REGION Network 1 (SCL)
   //---------------------------------------------------------------------
   //In this network first, we assign the ip address and port number for the printer (MarkemImaje). Then prepare the command for 
   //time synch, checking alarms, sending a batch number, intiating counter and selecting the label. one port for all data.
   //---------------------------------------------------------------------
   //
   REGION AddressAssign
       (*
       //Special case: if ip and port is entered correctly but still the communication not established, try onece more.
       IF #ConnectionStatus = False AND #ErrorIP = FALSE AND #ReTry = FALSE AND #ConnAgainT.Q = FALSE AND #TimeOutError = FALSE THEN
           #ReTry := True;
       ELSE
           #ReTry := FALSE;
       END_IF;
       *)
       // ip and port assign to the printer
       #Config := "LGF_StringToTaddr"(ipAddressString := #RemoteAddress, error => #ErrorIP, status => #StatusIP);
       //when IP address change, disconnect and connect again
       #ChangeIP_T(IN:=#RemoteAddressOld <> #RemoteAddress,
                   PT:=T#2S);
       IF #ChangeIP_T.Q OR #ErrorIP = TRUE THEN
           #IP_Change := TRUE;
       ELSE
           #IP_Change := FALSE;
       END_IF;
       #RemoteAddressOld := #RemoteAddress;
       FOR #i := 1 TO 4 DO
           #Configuration.connection.partnerIP.ADDR[#i] := USINT_TO_BYTE(#Config.REM_IP_ADDR[#i]);//assign ip address
       END_FOR;
       //assign id port and other setting for TCP communication
       #Configuration.connection.connectionID := #ID;
       #Configuration.connection.comService := 1;
       //if it is active connection
       IF #ConType = TRUE THEN
           #Configuration.connection.isClient := True;
           IF #Config.REM_PORT_NR = 0 THEN
               #Configuration.connection.partnerPort := 9100; // default port for Markem communication
           ELSE
               #Configuration.connection.partnerPort := #Config.REM_PORT_NR;
           END_IF;
       ELSE //if it is passive connection
           #Configuration.connection.isClient := FALSE;
           #Configuration.connection.localPort := 2000;
       END_IF;
   END_REGION
   REGION HMI
       // Data for the HMI
       #DatePrinted := DELETE(IN:=#Date, L:=2, P:=1);
       #TimePrinted := DELETE(IN := #Time, L := 2, P := 5);
       #TimePrinted := INSERT(IN1 := #TimePrinted, IN2 := ':', P := 2);
       IF #ExtDate <> '' THEN
           #ExpFlag := TRUE;
       ELSE
           #ExpFlag := FALSE;
       END_IF;
   END_REGION

   REGION Commands 
       // Creating Commands and preparing them to Send
       IF #Step = 1 THEN
           //command for time synchronisation
           #CommandHead := 'V21'; //head for time/date synch
           #SData[0] := #Start;
           Strg_TO_Chars(Strg := #CommandHead,
                         pChars := 1,
                         Cnt => #Dummy2,
                         Chars := #SData);
           #SData[4] := ' ';
           Strg_TO_Chars(Strg := #Date,
                         pChars := 0,
                         Cnt => #Dummy2,
                         Chars := #DateChar);
           FOR #i := 5 TO 8 DO
               #SData[#i] := #DateChar[#i - 5];
           END_FOR;
           #SData[9] := '-';
           #SData[10] := #DateChar[4];
           #SData[11] := #DateChar[5];
           #SData[12] := '-';
           #SData[13] := #DateChar[6];
           #SData[14] := #DateChar[7];
           #SData[15] := #NewLine;
           //sending time
           #SData[16] := #Start;
           #SData[17] := 'V';
           #SData[18] := '2';
           #SData[19] := '0';
           #SData[20] := ' ';
           Strg_TO_Chars(Strg := #Time,
                         pChars := 0,
                         Cnt => #Dummy2,
                         Chars := #TimeChar);
           #SData[21] := #TimeChar[0];
           #SData[22] := #TimeChar[1];
           #SData[23] := ':';
           #SData[24] := #TimeChar[2];
           #SData[25] := #TimeChar[3];
           #SData[26] := ':';
           #SData[27] := #TimeChar[4];
           #SData[28] := #TimeChar[5];
           #SData[29] := #End;
           #RLen := 2;
           #SLen := 30;
           #Step := 0;
           #STrig := TRUE;
           #RdataTime := TRUE;
           #RdataAlarm := FALSE;
           #RdataBatch := FALSE;
           #RdataMacro := FALSE;
       ELSIF #Step = 2 THEN
           //command for checking the alarms
           #CommandHead := 'S100'; //head for current status of the printer
           #SData[0] := #Start;
           Strg_TO_Chars(Strg := #CommandHead,
                         pChars := 1,
                         Cnt => #Dummy2,
                         Chars := #SData);
           #SData[5] := #End;
           #RLen := 34;
           #SLen := 6;
           #STrig := TRUE;
           #Step := 0;
           #RdataAlarm := TRUE;
           #RdataTime := FALSE;
           #RdataBatch := FALSE;
           #RdataMacro := FALSE;
       ELSIF #Step = 3 THEN
           //command for sending variable text
           #SData[0] := #Start;
           #CommandHead := 'W1 "';
           //GTIN number 14 digits
           Strg_TO_Chars(Strg := #CommandHead,
                         pChars := 1,
                         Cnt => #Dummy2,
                         Chars := #SData);
           Strg_TO_Chars(Strg := #GTIN_Number,
                         pChars := 5,
                         Cnt => #Dummy2,
                         Chars := #SData);
           #SData[19] := '"';
           #SData[20] := #NewLine;
           //Batch
           #CommandHead := '!W4 "';
           //Batch number 10 digits
           Strg_TO_Chars(Strg := #CommandHead,
                         pChars := 21,
                         Cnt => #Dummy2,
                         Chars := #SData);
           Strg_TO_Chars(Strg := #BatchNumber,
                         pChars := 26,
                         Cnt => #Dummy2,
                         Chars := #SData);
           #SData[36] := '"';
           #SData[37] := #NewLine;
           //Article number
           #CommandHead := '!W5 "';
           //Article number 10 digits
           Strg_TO_Chars(Strg := #CommandHead,
                         pChars := 38,
                         Cnt => #Dummy2,
                         Chars := #SData);
           Strg_TO_Chars(Strg := #ArtNumber,
                         pChars := 43,
                         Cnt => #Dummy2,
                         Chars := #SData);
           #SData[53] := '"';
           #SData[54] := #NewLine;
           //Ext date
           #CommandHead := '!W3 "';
           //Ext date 6 digits
           Strg_TO_Chars(Strg := #CommandHead,
                         pChars := 55,
                         Cnt => #Dummy2,
                         Chars := #SData);
           IF #ExtDate <> '' THEN //if expiration date is available 
               Strg_TO_Chars(Strg := #ExtDate,
                             pChars := 60,
                             Cnt => #Dummy2,
                             Chars := #SData);
           ELSE
               FOR #i := 60  TO 65 DO
                   #SData[#i] := ' ';
               END_FOR;
           END_IF;
           #SData[66] := '"';
           #SData[67] := #NewLine;
           //Machine ID
           #CommandHead := '!W6 "';
           //Machine ID 3 digits
           Strg_TO_Chars(Strg := #CommandHead,
                         pChars := 68,
                         Cnt => #Dummy2,
                         Chars := #SData);
           Strg_TO_Chars(Strg := #MachineID,
                         pChars := 73,
                         Cnt => #Dummy2,
                         Chars := #SData);
           //Reinit the counter 
           #SData[76] := '"';
           #SData[77] := #NewLine;
           VAL_STRG(IN := (#Serial+1),// +1 to make sure we have no TRP with same serial
                    SIZE := 0,
                    PREC := 0,
                    FORMAT := 0,
                    P := 1,
                    OUT => #SerialSTR);
           #SerialLen := LEN(#SerialSTR);
           #CommandHead := '!N1 ';//!N1 "Serial" 1 5 1
           Strg_TO_Chars(Strg := #CommandHead,
                         pChars := 78,
                         Cnt => #Dummy2,
                         Chars := #SData);
           #CommandHead := #SerialSTR;
           Strg_TO_Chars(Strg := #CommandHead,
                         pChars := 82,
                         Cnt => #Dummy2,
                         Chars := #SData);
           #CommandHead := ' 1 5 1';
           Strg_TO_Chars(Strg := #CommandHead,
                         pChars := 82+#SerialLen,
                         Cnt => #Dummy2,
                         Chars := #SData);
           #SData[82 + #SerialLen + 6] := #End;
           #RLen := 0;
           #SLen := INT_TO_UDINT( 82 + #SerialLen + 6 + 1);
           #Step := 0;
           #STrig := TRUE;
           #Selected := FALSE;
           #RdataTime := FALSE;
           #RdataAlarm := FALSE;
           #RdataBatch := TRUE;
           #RdataMacro := FALSE;
       //command for selectiong the Macro 
       ELSIF #Step = 4 THEN
           #CommandHead := 'M "'; //head for selecting the Macro
           #SData[0] := #Start;
           Strg_TO_Chars(Strg := #CommandHead,
                         pChars := 1,
                         Cnt => #Dummy2,
                         Chars := #SData);
           IF #ExtDate = '' THEN
               IF #Inverse = TRUE THEN
                   Strg_TO_Chars(Strg := #LabelNameInv,
                                 pChars := 4,
                                 Cnt => #Dummy2,
                                 Chars := #SData);
               ELSE
                   Strg_TO_Chars(Strg := #LabelName,
                                 pChars := 4,
                                 Cnt => #Dummy2,
                                 Chars := #SData);
               END_IF;
           ELSE
               IF #Inverse = TRUE THEN
                   Strg_TO_Chars(Strg := #LabelNameExpInv,
                                 pChars := 4,
                                 Cnt => #Dummy2,
                                 Chars := #SData);
               ELSE
                   Strg_TO_Chars(Strg := #LabelNameExp,
                                 pChars := 4,
                                 Cnt => #Dummy2,
                                 Chars := #SData);
               END_IF;
           END_IF;
           #SData[16] := '"';
           #SData[17] := #NewLine;
           IF #Stop = TRUE THEN
               #SData[18] := ' ';
               #SData[19] := 'p';
           ELSE
               #SData[18] := #Start;
               #SData[19] := 'p';
           END_IF;
           #SData[20] := #End;
           #RLen := 2;
           #SLen := 21;
           #Step := 0;
           #STrig := TRUE;
           #RdataTime := FALSE;
           #RdataAlarm := FALSE;
           #RdataBatch := FALSE;
           #RdataMacro := TRUE;
       ELSE
           #STrig := FALSE;
       END_IF;
   END_REGION

   REGION Feedback
       // Statement section REGION
       //Expect to receive "ACT"
       IF #DataReceived = TRUE THEN
           #StartTNR := FALSE;
           IF #RdataTime = TRUE THEN //check for the feedback for the time command
               FOR #i := 0 TO 56 DO
                   #TimeReceivedData[#i] := #RData[#i];
               END_FOR;
               IF #TimeReceivedData[0] = #NewLine THEN
                   #TimeOK := TRUE;
                   #TimeReceivedData[0] := 16#30;//clear the buffer
               ELSE
                   #TimeOK := FALSE;
               END_IF;
               #RdataTime := FALSE; // make the flag false
           ELSIF #RdataAlarm = TRUE THEN//check for the feedback for the alarm command
               FOR #i := 0 TO 56 DO
                   #AlarmReceivedData[#i] := #RData[#i];
               END_FOR;
               IF #AlarmReceivedData[32] = #End THEN // the plc receives the responce
                   #AlarmCheck := TRUE;
                   #AlarmReceivedData[32] := 16#30;//clear the buffer
                   FOR #i := 0 TO 31 DO//save the status data for processing
                       IF #AlarmReceivedData[#i] = '1' THEN
                           #PrinterAlarmStatus[#i] := TRUE;
                       ELSE
                           #PrinterAlarmStatus[#i] := FALSE;
                       END_IF;
                   END_FOR;
               ELSE
                   #AlarmCheck := FALSE;
               END_IF;
               #RdataAlarm := FALSE;
           //ELSIF #RdataBatch = TRUE THEN //no feedback from the command except batch
               //         FOR #i := 0 TO 56 DO
               //            #BatchReceivedData[#i] := #RData[#i];
               //        END_FOR;
               //       IF #BatchReceivedData[0] = 16#24 THEN
             //  #BatchOK := TRUE;
               //           #BatchReceivedData[0] := 16#30;//clear the buffer
               //       ELSE
               //        #BatchOK := FALSE;
               //    END_IF;
               //     #RdataBatch := FALSE;
           ELSIF #RdataMacro = TRUE OR #RdataBatch = TRUE THEN
               FOR #i := 0 TO 56 DO
                   #MacroReceivedData[#i] := #RData[#i];
               END_FOR;
               IF #MacroReceivedData[0] = #NewLine THEN // the plc receives the responce
                   #LabelOK := TRUE;
                   #MacroReceivedData[0] := 16#30;//clear the buffer
               ELSE
                   #LabelOK := FALSE;
               END_IF;
               #RdataMacro := FALSE;
           END_IF;
       ELSIF #DataSent = TRUE AND #RdataAlarm = TRUE OR #RdataTime = TRUE OR #RdataMacro = TRUE THEN // command send noting received
           #StartTNR := TRUE;
           IF #RdataTime = TRUE THEN
               #TimeOK := FALSE;
           END_IF;
           IF #RdataAlarm = TRUE THEN
               #AlarmCheck := FALSE;
           END_IF;
           IF #RdataMacro = TRUE THEN
               #LabelOK := FALSE;
           END_IF;
       END_IF;
   END_REGION

   REGION Sending
       //selecting the label properties for every instalation of the new printer or power OFF then ON
       #SelectingR(CLK:=#LabelSelecting);
       #ReconnectR(CLK := #ConnectionStatus);
       #InverseR(CLK:=#Inverse);
       #InverseF(CLK:=#Inverse);
        // it is assumed at every reconnection the label is gone so, we send it again
       IF #SelectingR.Q = TRUE OR #ReconnectR.Q = TRUE OR #InverseR.Q = TRUE OR #InverseF.Q = TRUE THEN
           #Step := 4;
           #Selected := TRUE;
       END_IF;
       // set the step to 3 after label is selecting (small delay to make sure that the label is loaded)
       #BatchAfterLabelT(IN := #Selected,
                         PT := T#5S);
       IF #BatchAfterLabelT.Q = TRUE THEN
           #Step := 3;
       END_IF;
       // Send the updateble data when it is changed and step 4 is done
       IF #PlainDataChanged = TRUE AND #SelectingR.Q = FALSE THEN
           #Step := 3;
           #Selected := FALSE;
       END_IF;
       // Send time and alarm commands
       //every 10 minute synchronise time
       #TimeSynchT(IN := #TimeSynchEnable,
                  PT := #TimeSynchPeriod);
       IF #TimeSynchT.Q = TRUE THEN
           #Step := 1;
           #TimeSynchEnable := FALSE;
       ELSIF #ConnectionStatus = TRUE AND NOT (#SelectingR.Q = TRUE OR #ReconnectR.Q = TRUE OR #InverseR.Q = TRUE OR #InverseF.Q = TRUE) AND #PlainDataChanged = FALSE THEN
           #TimeSynchEnable := True;
       ELSE
           #TimeSynchEnable := FALSE;
       END_IF;
       //every 5 minute check for alarm
       #AlarmCheckT(IN := #AlarmCheckEnable,
                   PT := #AlarmCheckPeriod + T#20MS);//+20ms to avoid conflict
       IF #AlarmCheckT.Q = TRUE THEN
           #Step := 2;
           #AlarmCheckEnable := FALSE;
       ELSIF #ConnectionStatus = TRUE AND NOT (#SelectingR.Q = TRUE OR #ReconnectR.Q = TRUE OR #InverseR.Q = TRUE OR #InverseF.Q = TRUE) AND #PlainDataChanged = FALSE THEN
           #AlarmCheckEnable := TRUE;
       ELSE
           #AlarmCheckEnable := FALSE;
       END_IF;
   END_REGION
   (*
   REGION ConnReestablised
       // connection Re-Established Rotinue. It try 5 times to connect to the printer, if not succsess enable time out error
       #ConnAgainT(IN := #ReTry,
                  PT := T#5S);// time out for reconnection
       //try five times to connect
       #ConnTryCountC(CU := #ReTry,
                     R := #ConnectionStatus,
                     PV := 5,
                     Q => #TimeOutError);
   END_REGION
   *)
   REGION send try
       //if not receiving feedback after 10ms send a commad again
       #NotReceiveT(IN := #StartTNR,
                   PT := #TimeNR,
                   Q => #SendAgainTrigger);
       IF #SendAgainTrigger = TRUE THEN
           #StartTNR := FALSE;
       END_IF;
    //   #NotReceivingError(IN:= NOT(#TimeOK AND #LabelOK AND #NoAlarm = FALSE), // if we are not receiving a feedback after sending two times pop up an alarm
    //                      PT:=T#90S,
    //                      Q=>#CommandError);
   END_REGION

   REGION Counter
       // count the number of the trigger and initiated it when sending the label information. the counter only restarted when the batch changed. 
       #ExtTriggerR(CLK:=#ExtTrigger);
       IF #ExtTriggerR.Q = TRUE THEN
           "Counter_32Bit_1"(Varia := 1,
                           CountedValue := #Serial);
       END_IF;
       IF #Serial > 99999 OR #PlainDataChanged = TRUE THEN //restart the counter if it reaches the limit or data changed at Plain
           #Serial := 0;
       END_IF;
   END_REGION
END_REGION
END_FUNCTION_BLOCK

FUNCTION_BLOCK "Domino_AX"   // FB6, LAD
{ S7_Optimized_Access := 'TRUE' }
VERSION : 0.1
   VAR_INPUT
      RemoteAddress : String[20];
      ConnectionStatus : Bool;
      ID : Conn_Ouc;
      ConType : Bool;
      ArtFlag : Bool;
      MDR_Flag : Bool;
      BatchStatus : USInt;
      BatchNumber : String;
      ArtBaseNumber : String;
      MarketRegCode : String;
      ExtDate : String;
      "Date" : String;
      "Time" : String;
      PlainDataChanged : Bool;
      DataReceived : Bool;
      DataReceivedBatch : Bool;
      DataSent : Bool;
      DataSentBatch : Bool;
      TimeSynchPeriod : Time := T#10M;
      AlarmCheckPeriod : Time := T#5M;
      RDataBatch : Array[0..56] of Byte;
      RData : Array[0..56] of Byte;
      NMDR_LabelName : String;
      LabelSelecting : Bool;
   END_VAR
   VAR_OUTPUT
      ErrorIP : Bool;
      BatchOK : Bool;
      AlarmCheck : Bool;
      TimeOK : Bool;
      LabelOK : Bool;
   END_VAR
   VAR
      Config : TADDR_Param;
      Configuration : "typeLCom_Config";
      ConfigurationBatch : "typeLCom_Config";
      RLen : UDInt;
      RLenMDR : UDInt;
      SLen : UDInt;
      SLenMDR : UDInt;
      SData : Array[0..56] of Byte;
      SDataMDR : Array[0..99] of Byte;
      StartTNRMDR : Bool;
      StartTNR : Bool;
      TimeNR : Time := T#1m;
      SendAgainTrigger : Bool;
      SendAgainTriggerBatch : Bool;
      NotReceiveT : TON_TIME;
      NotReceiveBatchT : TON_TIME;
      TimeSynchEnable : Bool := false;
      TimeSynchT : TON_TIME;
      AlarmCheckEnable : Bool := false;
      AlarmCheckT : TON_TIME;
      STrig : Bool;
      StrigBatch : Bool;
      "Step" : UDInt;
      AlarmReceivedData : Array[0..56] of Byte;
      TimeReceivedData : Array[0..56] of Byte;
      BatchReceivedData : Array[0..56] of Byte;
      LabelReceivedData : Array[0..56] of Byte;
      PrinterAlarmStatus : Array[0..8] of Char;
      RdataTime : Bool;
      RdataAlarm : Bool;
      RdataLabel : Bool;
      BlockedProduct : Bool;
      SelectingR : R_TRIG;
      Selected : Bool;
      ReconnectR : R_TRIG;
      MDR_R : R_TRIG;
      MDR_F : F_TRIG;
      BlockedR : R_TRIG;
      BlockedF : F_TRIG;
      ActualNMDR_Label : String;
      NLabelChanged : Bool;
      BatchAfterLabelT : TON_TIME;
      ChangeIP_T : TP_TIME;
      IP_Change : Bool;
      RemoteAddressOld : String;
   END_VAR
   VAR_TEMP
      StatusIP : Word;
      Dummy2 : UInt;
      i : Int;
      CommandHead : String;
      SecondRowSTR : String;
      SecondRowSTR1 : String;
      LenDummy : Int;
      ArtLen : Int;
      LenLabel : Int;
      LenLabelSTR : String;
      LabelCommand : String;
   END_VAR
   VAR CONSTANT
      Start : Char := '$1B';
      Start1 : Char := '$02';
      End1 : Char := '$03';
      End : Char := '$04';
      MDR_LabelName1 : String := 'MDR1';
      MDR_LabelName2 : String := 'MDR2';
   END_VAR
BEGIN

REGION Network 1 (SCL)
   //---------------------------------------------------------------------
   //In this network first, we assign the ip address and port number for the printer (Domino_AX). Then prepare the command for 
   //time synch, receiving alarms and sending a batch number. one port (16000) for the batch number and another port for the rest.
   //---------------------------------------------------------------------
   REGION Address_Assign
       (*
       //Special case: if ip and port is entered correctly but still the communication not established, try onece more.
       IF #ConnectionStatus = False AND #ErrorIP = FALSE AND #ReTry = FALSE AND #ConnAgainT.Q = FALSE AND #TimeOutError = FALSE THEN
           #ReTry := True;
       ELSE
           #ReTry := FALSE;
       END_IF;
       *)
       // ip and port assign to the printer
       #Config := "LGF_StringToTaddr"(ipAddressString := #RemoteAddress, error => #ErrorIP, status => #StatusIP);
       //when IP address change, disconnect and connect again
       #ChangeIP_T(IN := #RemoteAddressOld <> #RemoteAddress,
                   PT := T#2S);
       IF #ChangeIP_T.Q OR #ErrorIP = TRUE THEN
           #IP_Change := TRUE;
       ELSE
           #IP_Change := FALSE;
       END_IF;
       #RemoteAddressOld := #RemoteAddress;
       FOR #i := 1 TO 4 DO
          #Configuration.connection.partnerIP.ADDR[#i] := USINT_TO_BYTE(#Config.REM_IP_ADDR[#i]);//assign ip address
          #ConfigurationBatch.connection.partnerIP.ADDR[#i] := USINT_TO_BYTE(#Config.REM_IP_ADDR[#i]);//assign ip address
      END_FOR;

       //assign id port and other setting for TCP communication
       #Configuration.connection.connectionID := #ID;
       #Configuration.connection.comService := 1;
       #ConfigurationBatch.connection.connectionID := #ID + 1;
       #ConfigurationBatch.connection.comService := 1;
       #ConfigurationBatch.connection.isClient := True;
       #ConfigurationBatch.connection.partnerPort := 16000;// only for domino printer
         //if it is active connection
       IF #ConType = TRUE THEN
           #Configuration.connection.isClient := True;
           IF #Config.REM_PORT_NR = 0 THEN
               #Configuration.connection.partnerPort := 7000; // default port for domino communication
           ELSE
               #Configuration.connection.partnerPort := #Config.REM_PORT_NR;
           END_IF;
       ELSE //if it is passive connection
           #Configuration.connection.isClient := FALSE;
           #Configuration.connection.localPort := 2000;
       END_IF;

   END_REGION
   REGION Trigger
       // Trigger signal to send a correct data for print when Batch ended
       IF #BatchStatus = 3 THEN
           #BlockedProduct := TRUE;
       ELSE
           #BlockedProduct := FALSE;
       END_IF;
       // Trigger signal to send Non-MDR label when it is changed from the screen
       IF #MDR_Flag = FALSE AND #ActualNMDR_Label <> #NMDR_LabelName THEN
           #NLabelChanged := TRUE;
           #ActualNMDR_Label := #NMDR_LabelName;
       ELSE
           #NLabelChanged := FALSE;
       END_IF;
   END_REGION

   REGION Commands
         //command for time synchronisation
         IF #Step = 1 THEN
             #CommandHead := 'C'; //head for time
             #SData[0] := #Start;
             Strg_TO_Chars(Strg := #CommandHead,
                           pChars := 1,
                           Cnt => #Dummy2,
                           Chars := #SData);
             Strg_TO_Chars(Strg := #Date,
                           pChars := 2,
                           Cnt => #Dummy2,
                           Chars := #SData);
             #SData[10] := '0';
             #SData[11] := '0';
             Strg_TO_Chars(Strg := #Time,
                           pChars := 12,
                           Cnt => #Dummy2,
                           Chars := #SData);
             #SData[18] := #End;
             #RLen := 1;
             #SLen := 19;
             #STrig := TRUE;
             #Step := 0; //idea state
             #RdataTime := TRUE;
             #RdataAlarm := FALSE;
             #RdataLabel := FALSE;

         ELSIF #Step = 2 THEN
             //command for checking the alarms
             #CommandHead := 'O1?'; //head for current status of the printer
             #SData[0] := #Start;
             Strg_TO_Chars(Strg := #CommandHead,
                           pChars := 1,
                           Cnt => #Dummy2,
                           Chars := #SData);
             #SData[4] := #End;
             #RLen := 9;
             #SLen := 5;
             #STrig := TRUE;
             #Step := 0; 
             #RdataAlarm := TRUE;
             #RdataTime := FALSE;
             #RdataLabel := FALSE;
             (*  we should creat a MDR layout at the Printer with two fields. one id used for batch+art base and the 
                   second is use for market Reg and Ext date*)
                   //Constructiong the buffer command in the first row
         ELSIF #Step=3 THEN
             #RLenMDR := 1; // receive 0x06 as an acknowledgment
             #StrigBatch := TRUE;
             #Step := 0;
             #Selected := FALSE;
                 #SDataMDR[0] := #Start1;
                 Strg_TO_Chars(Strg := #BatchNumber,
                               pChars := 1,
                               Cnt => #Dummy2,
                               Chars := #SDataMDR);
                 IF #ArtFlag = TRUE AND #MarketRegCode <> '' AND #ExtDate <> '' THEN // print all information in two rows
                     #SDataMDR[11] := ' '; //space
                     #SDataMDR[12] := 'A';
                     #SDataMDR[13] := 'R';
                     #SDataMDR[14] := 'T';
                     #ArtLen := LEN(#ArtBaseNumber);
                     Strg_TO_Chars(Strg := #ArtBaseNumber,
                                   pChars := 15,
                                   Cnt => #Dummy2,
                                   Chars := #SDataMDR);
                     IF #BatchStatus = 3 THEN //add a sign '+' at the con
                         #SDataMDR[15 + #ArtLen] := '+';

                     ELSE
                         #SDataMDR[15 + #ArtLen] := ' ';
                     END_IF;
                     #SDataMDR[15 + #ArtLen + 1] := ',';//seprator for the second row
                     #SecondRowSTR := CONCAT(IN1 := #MarketRegCode, IN2 := 'BBD');
                     #SecondRowSTR1 := CONCAT(IN1 := #SecondRowSTR, IN2 := #ExtDate);
                     #LenDummy := LEN(#SecondRowSTR1);
                     Strg_TO_Chars(Strg := #SecondRowSTR1,
                                   pChars := 15 + #ArtLen + 2,
                                   Cnt => #Dummy2,
                                   Chars := #SDataMDR);
                     #SDataMDR[15 + #ArtLen + 2 + #LenDummy] := #End1;
                     #SLenMDR := 15 + #ArtLen + 2 + #LenDummy + 1;
                 ELSIF #ArtFlag = TRUE AND #MarketRegCode <> '' AND #ExtDate = '' THEN // print all information exept expiration date in two rows
                     #SDataMDR[11] := ' '; //space
                     #SDataMDR[12] := 'A';
                     #SDataMDR[13] := 'R';
                     #SDataMDR[14] := 'T';
                     #ArtLen := LEN(#ArtBaseNumber);
                     Strg_TO_Chars(Strg := #ArtBaseNumber,
                                   pChars := 15,
                                   Cnt => #Dummy2,
                                   Chars := #SDataMDR);
                     IF #BatchStatus = 3 THEN //add a sign '+' at the con
                         #SDataMDR[15 + #ArtLen] := '+';

                     ELSE
                         #SDataMDR[15 + #ArtLen] := ' ';
                     END_IF;
                     #SDataMDR[15 + #ArtLen + 1] := ',';//seprator for the second row
                     #LenDummy := LEN(#MarketRegCode);
                     Strg_TO_Chars(Strg := #MarketRegCode,
                                   pChars := 15 + #ArtLen + 2,
                                   Cnt => #Dummy2,
                                   Chars := #SDataMDR);
                     #SDataMDR[15 + #ArtLen + 2 + #LenDummy] := #End1;
                     #SLenMDR := 15 + #ArtLen + 2 + #LenDummy + 1;
                 ELSIF #ArtFlag = TRUE AND #MarketRegCode = '' AND #ExtDate <> '' THEN // print all information exept Market reg code in two rows
                     #SDataMDR[11] := ' '; //space
                     #SDataMDR[12] := 'A';
                     #SDataMDR[13] := 'R';
                     #SDataMDR[14] := 'T';
                     #ArtLen := LEN(#ArtBaseNumber);
                     Strg_TO_Chars(Strg := #ArtBaseNumber,
                                   pChars := 15,
                                   Cnt => #Dummy2,
                                   Chars := #SDataMDR);
                     IF #BatchStatus = 3 THEN //add a sign '+' at the con
                         #SDataMDR[15 + #ArtLen] := '+';

                     ELSE
                         #SDataMDR[15 + #ArtLen] := ' ';
                     END_IF;
                     #SDataMDR[15 + #ArtLen + 1] := ',';//seprator for the second row
                     #SecondRowSTR1 := CONCAT(IN1 := 'BBD', IN2 := #ExtDate);
                     #LenDummy := LEN(#SecondRowSTR1);
                     Strg_TO_Chars(Strg := #SecondRowSTR1,
                                   pChars := 15 + #ArtLen + 2,
                                   Cnt => #Dummy2,
                                   Chars := #SDataMDR);
                     #SDataMDR[15 + #ArtLen + 2 + #LenDummy] := #End1;
                     #SLenMDR := 15 + #ArtLen + 2 + #LenDummy + 1;
                 ELSIF #ArtFlag = TRUE AND #MarketRegCode = '' AND #ExtDate = '' THEN // print only in one row
                     #SDataMDR[11] := ' '; //space
                     #SDataMDR[12] := 'A';
                     #SDataMDR[13] := 'R';
                     #SDataMDR[14] := 'T';
                     #ArtLen := LEN(#ArtBaseNumber);
                     Strg_TO_Chars(Strg := #ArtBaseNumber,
                                   pChars := 15,
                                   Cnt => #Dummy2,
                                   Chars := #SDataMDR);
                     IF #BatchStatus = 3 THEN //add a sign '+' at the con
                         #SDataMDR[15 + #ArtLen] := '+';

                     ELSE
                         #SDataMDR[15 + #ArtLen] := ' ';
                     END_IF;
                     #SDataMDR[16 + #ArtLen] := #End1;
                     #SLenMDR := 16 + #ArtLen + 1;
                 ELSIF #ArtFlag = FALSE AND #MarketRegCode <> '' AND #ExtDate <> '' THEN // print all information exept art flag  in two rows
                     IF #BatchStatus = 3 THEN //add a sign '+' at the con
                         #SDataMDR[11] := '+';

                     ELSE
                         #SDataMDR[11] := ' ';
                     END_IF;
                     #SDataMDR[12] := ',';//seprator for the second row
                     #SecondRowSTR := CONCAT(IN1 := #MarketRegCode, IN2 := 'BBD');
                     #SecondRowSTR1 := CONCAT(IN1 := #SecondRowSTR, IN2 := #ExtDate);
                     #LenDummy := LEN(#SecondRowSTR1);
                     Strg_TO_Chars(Strg := #SecondRowSTR1,
                                   pChars := 13,
                                   Cnt => #Dummy2,
                                   Chars := #SDataMDR);
                     #SDataMDR[13 + #LenDummy] := #End1;
                     #SLenMDR := 13 + #LenDummy + 1;
                 ELSIF #ArtFlag = FALSE AND #MarketRegCode <> '' AND #ExtDate = '' THEN // print all information exept expiration art number and ext date in two rows
                     IF #BatchStatus = 3 THEN //add a sign '+' at the con
                         #SDataMDR[11] := '+';

                     ELSE
                         #SDataMDR[11] := ' ';
                     END_IF;
                     #SDataMDR[12] := ',';//seprator for the second row
                     #LenDummy := LEN(#MarketRegCode);
                     Strg_TO_Chars(Strg := #MarketRegCode,
                                   pChars := 13,
                                   Cnt => #Dummy2,
                                   Chars := #SDataMDR);
                     #SDataMDR[13 + #LenDummy] := #End1;
                     #SLenMDR := 13 + #LenDummy + 1;
                 ELSIF #ArtFlag = FALSE AND #MarketRegCode = '' AND #ExtDate <> '' THEN // print in one row
                     IF #BatchStatus = 3 THEN //add a sign '+' at the con
                         #SDataMDR[11] := '+';

                     ELSE
                         #SDataMDR[11] := ' ';
                     END_IF;
                     #SDataMDR[12] := ',';//seprator for the second row
                     #SecondRowSTR1 := CONCAT(IN1 := 'BBD', IN2 := #ExtDate);
                     #LenDummy := LEN(#SecondRowSTR1);
                     Strg_TO_Chars(Strg := #SecondRowSTR1,
                                   pChars := 13,
                                   Cnt => #Dummy2,
                                   Chars := #SDataMDR);
                     #SDataMDR[13 + #LenDummy] := #End1;
                     #SLenMDR := 13 + #LenDummy + 1;
                 ELSE // print only batch
                     IF #BatchStatus = 3 THEN //add a sign '+' at the con
                         #SDataMDR[11] := '+';

                     ELSE
                         #SDataMDR[11] := ' ';
                     END_IF;
                     #SDataMDR[12] := #End1;
                     #SLenMDR := 13;
                 END_IF;
         ELSIF #Step =4 THEN
             //command for selecting the label
             #CommandHead := 'ON1'; //head for current status of the printer
             #SData[0] := #Start;
             Strg_TO_Chars(Strg := #CommandHead,
                           pChars := 1,
                           Cnt => #Dummy2,
                           Chars := #SData);
             IF #MDR_Flag = TRUE THEN //select the MDR layout 
                 IF #ExtDate <> '' OR #MarketRegCode <> '' THEN
                     #LabelCommand := CONCAT(IN1 := '04', IN2 := #MDR_LabelName2);
                 ELSE
                     #LabelCommand := CONCAT(IN1 := '04', IN2 := #MDR_LabelName1);
                 END_IF;
                 Strg_TO_Chars(Strg := #LabelCommand,
                               pChars := 4,
                               Cnt => #Dummy2,
                               Chars := #SData);
                 #SData[10] := #End;
                 #RLen := 1;
                 #SLen := 11;
             ELSE
                 #LenLabel := LEN(#NMDR_LabelName);
                 VAL_STRG(IN := #LenLabel,
                          SIZE := 2,
                          PREC := 0,
                          FORMAT := 0,
                          P := 1,
                          OUT => #LenLabelSTR);
                 #LabelCommand := CONCAT(IN1 := #LenLabelSTR, IN2 := #NMDR_LabelName);

                 Strg_TO_Chars(Strg := #LabelCommand,
                               pChars := 4,
                               Cnt => #Dummy2,
                               Chars := #SData);
                 FOR #i := 4 TO 5 DO //check for null char due to size
                     IF #SData[#i] = ' ' THEN
                         #SData[#i] := '0';
                     END_IF;
                 END_FOR;
                 #SData[6 + #LenLabel] := #End;
                 #RLen := 1;
                 #SLen := 7 + #LenLabel;
             END_IF;
             #STrig := TRUE;
             #Step := 0; 
             #RdataAlarm := FALSE;
             #RdataTime := FALSE;
             #RdataLabel := TRUE;
         ELSE
             #STrig := FALSE;
             #StrigBatch := FALSE;
         END_IF;
     END_REGION
       REGION Feedback
           // Statement section REGION
           //Expect to receive "ACT"
           IF #DataReceived = TRUE THEN
               #StartTNR := FALSE;
               IF #RdataTime = TRUE THEN //check for the feedback for the time command
                   FOR #i := 0 TO 56 DO
                       #TimeReceivedData[#i] := #RData[#i];
                   END_FOR;
                   IF #TimeReceivedData[0] = 16#06 THEN
                       #TimeOK := TRUE;
                       #TimeReceivedData[0] := 16#30;//clear the buffer
                   ELSE
                       #TimeOK := FALSE;
                   END_IF;
                   #RdataTime := FALSE;

               ELSIF #RdataAlarm = TRUE THEN//check for the feedback for the alarm command
                   FOR #i := 0 TO 56 DO
                       #AlarmReceivedData[#i] := #RData[#i];
                   END_FOR;
                   IF #AlarmReceivedData[1] = 'O' AND #AlarmReceivedData[2] = '1' THEN // check the responce and save them
                       #AlarmCheck := TRUE;
                       FOR #i := 0 TO 8 DO
                           #PrinterAlarmStatus[#i] := #AlarmReceivedData[#i];//save the status data for processing
                       END_FOR;
                       #AlarmReceivedData[1] := '0';//clear the buffer
                   ELSE
                       #AlarmCheck := FALSE;
                   END_IF;
                   #RdataAlarm := FALSE;
               ELSIF #RdataLabel = TRUE THEN // check for the label command feedback
                   FOR #i := 0 TO 56 DO
                       #LabelReceivedData[#i] := #RData[#i];
                   END_FOR;
                   IF #LabelReceivedData[0] = 16#06 THEN // check the responce and save them
                       #LabelOK := TRUE;
                       #LabelReceivedData[0] := '0';//clear the buffer
                   ELSE
                       #LabelOK := FALSE;
                   END_IF;
                   #RdataLabel := FALSE;
               END_IF;
           ELSIF #DataSent = TRUE THEN // command send noting received
                   #StartTNR := TRUE;
                   IF #RdataTime = TRUE THEN
                       #TimeOK := FALSE;
                   END_IF;
                   IF #RdataAlarm = TRUE THEN
                       #AlarmCheck := FALSE;
                   END_IF;
                   IF #RdataLabel = TRUE THEN
                       #LabelOK := FALSE;
                   END_IF;
               END_IF;
               //Expect to receive "ACT" for external Info Command
               IF #DataReceivedBatch = TRUE THEN
                   #StartTNRMDR := FALSE;
                   FOR #i := 0 TO 56 DO
                       #BatchReceivedData[#i] := #RDataBatch[#i];
                   END_FOR;
                   IF #BatchReceivedData[0] = 16#06 THEN
                       #BatchOK := TRUE;
                   ELSE
                       #BatchOK := FALSE;
                   END_IF;
               ELSIF #DataSentBatch = TRUE THEN // command send noting received
                   #BatchOK := FALSE;
                   #StartTNRMDR := TRUE;
               END_IF;
       END_REGION

       REGION Sending
     // Send time, alarm and label commands
           #SelectingR(CLK:=#LabelSelecting);
           #ReconnectR(CLK:=#ConnectionStatus);
           #MDR_R(CLK := #MDR_Flag);
           #MDR_F(CLK:=#MDR_Flag);
           #BlockedR(CLK:=#BlockedProduct);
           #BlockedF(CLK:=#BlockedProduct);
           //select the label
           IF #MDR_F.Q= TRUE OR #MDR_R.Q =TRUE OR #SelectingR.Q = TRUE OR #ReconnectR.Q = TRUE OR #NLabelChanged = TRUE THEN
               #Step := 4; //selecting the label
               IF #MDR_Flag = TRUE THEN
                   #Selected := TRUE;
               END_IF;
           END_IF;
           // set the step to 3 after label is selected (small delay to make sure that the label is loaded)
           #BatchAfterLabelT(IN := #Selected,
                             PT := T#10S);
           IF #BatchAfterLabelT.Q = TRUE THEN
               #Step := 3;
           END_IF;
           //send the update information
           // Send the updatable data when it is changed and step 4 is done
           IF (#PlainDataChanged = TRUE OR #BlockedR.Q = TRUE OR #BlockedF.Q = TRUE) AND #SelectingR.Q = FALSE THEN
               #Step := 3; //send plain data
               #Selected := FALSE;
           END_IF;
     // synchronize time
    #TimeSynchT(IN:=#TimeSynchEnable,
               PT:=#TimeSynchPeriod);
    IF #TimeSynchT.Q = TRUE THEN
        #Step := 1;
        #TimeSynchEnable := FALSE;
    ELSIF #ConnectionStatus = TRUE AND NOT (#MDR_F.Q= TRUE OR #MDR_R.Q =TRUE OR #SelectingR.Q = TRUE OR #ReconnectR.Q = TRUE OR #NLabelChanged = TRUE) AND NOT (#PlainDataChanged = TRUE OR #BlockedR.Q = TRUE OR #BlockedF.Q = TRUE) THEN
        #TimeSynchEnable := TRUE;
    ELSE
        #TimeSynchEnable := FALSE;
    END_IF;
      // check the alarm
    #AlarmCheckT(IN:=#AlarmCheckEnable,
                PT:=#AlarmCheckPeriod+T#20MS);//+20ms to avoid conflict
    IF #AlarmCheckT.Q = TRUE THEN
        #Step := 2;
        #AlarmCheckEnable := FALSE;
    ELSIF #ConnectionStatus = TRUE AND NOT (#MDR_F.Q= TRUE OR #MDR_R.Q =TRUE OR #SelectingR.Q = TRUE OR #ReconnectR.Q = TRUE OR #NLabelChanged = TRUE) AND NOT (#PlainDataChanged = TRUE OR #BlockedR.Q = TRUE OR #BlockedF.Q = TRUE) THEN
        #AlarmCheckEnable := TRUE;
    ELSE
        #AlarmCheckEnable := FALSE;
    END_IF;
   END_REGION
    REGION send try
         //if not receiving feedback after 10ms send a commad again
         #NotReceiveT(IN := #StartTNR,
                     PT := #TimeNR,
                     Q => #SendAgainTrigger);
         #NotReceiveBatchT(IN := #StartTNRMDR,
                          PT := #TimeNR,
                          Q => #SendAgainTriggerBatch);
         IF #SendAgainTrigger = TRUE THEN
             #StartTNR := FALSE;
         END_IF;
         IF #SendAgainTriggerBatch = TRUE THEN
             #StartTNRMDR := FALSE;
         END_IF;
     END_REGION
     (*
     REGION ConnReestablised
         // connection Re-Established Rotinue. It try 5 times to connect to the printer, if not succsess enable time out error
         #ConnAgainT(IN := #ReTry,
                     PT := T#5S);// time out for reconnection
         //try five times to connect
         #ConnTryCountC(CU := #ReTry,
                       R := #ConnectionStatus,
                       PV := 5,
                       Q => #TimeOutError);
     END_REGION
     *)
END_REGION
END_FUNCTION_BLOCK

FUNCTION_BLOCK "ErrorHandeling"   // FB8, LAD
{ S7_Optimized_Access := 'TRUE' }
VERSION : 0.1
BEGIN
END_FUNCTION_BLOCK

FUNCTION_BLOCK "Counter_32Bit"   // FB9, FBD
{ S7_Optimized_Access := 'TRUE' }
AUTHOR : GeLa
VERSION : 0.1
   VAR_INPUT
      VARIA : DInt;
   END_VAR
   VAR_IN_OUT
      COUNTED_VALUE : DWord;
   END_VAR
   VAR
      COUNTED_VALUE_TMP1 : DInt;
   END_VAR
BEGIN

REGION Network 1
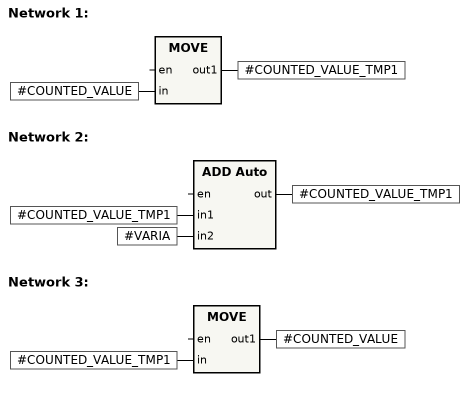
   #COUNTED_VALUE_TMP1 := #COUNTED_VALUE;
END_REGION

REGION Network 2
   #COUNTED_VALUE_TMP1 := #COUNTED_VALUE_TMP1 + #VARIA;
END_REGION

REGION Network 3
   #COUNTED_VALUE := #COUNTED_VALUE_TMP1;
END_REGION
END_FUNCTION_BLOCK

FUNCTION_BLOCK "TRP"   // FB10, FBD
{ S7_Optimized_Access := 'TRUE' }
VERSION : 0.1
   VAR
      edge : Array[0..15] of Bool;
      edge1 : Bool;
      edge2 : Bool;
      MDRTlac : Bool;
      OPC_HandleTRP_Instance : "TRP_PlainHandle";
      MarkemImaje : "MarkemImaje_2200";
      CommandSending_Markem : "LCom_Communication";
      Reader_2D_Instance : "Reader_2D";
      ReaderVerification_Instance : "ReaderVerification";
      TRP_PrinterStatus_Instance : "TRP_PrinterStatus";
   END_VAR
   VAR_TEMP
      tmp : Word;
      tmp_u : UInt;
   END_VAR
   VAR_TEMP   // added for the SCL form of the ladder/FBD networks
      _w1 : Bool;
      _w2 : Bool;
      _w3 : Bool;
      _w4 : Bool;
   END_VAR
BEGIN

REGION Network 2